                       IF "time_compare"(time_1 := #expire_date_time, time_2 := #current_time, difference_treshold := LT#0s) = true THEN

                           #shaker_batch_code_str[#runtime_shaker_index_finding_Instance.shaker_index - 1] := #batch_no;

                           IF #chemical = "DB_chemical_code".Application_bottle_code_Primer_DV954V1 THEN
                               #shaker_chemical_type_str[#runtime_shaker_index_finding_Instance.shaker_index - 1] := 'Primer DV 954 V1';
                               #shaker_door_lock_control_Instance.mixer_door_lock_enable[#runtime_shaker_index_finding_Instance.shaker_index - 1] := true;
                               #label_scanned := false;
                           ELSIF #chemical = "DB_chemical_code".Application_bottle_code_Primer_SIKA_207 THEN
                               #shaker_chemical_type_str[4] := 'Primer SIKA 207';
                               #shaker_door_lock_control_Instance.mixer_door_lock_enable[4] := true;
                               #label_scanned := false;
                           ELSE
                               #error_state := 256;
                               #shake_deinit := true;
                               #shaker_batch_code_str[#runtime_shaker_index_finding_Instance.shaker_index - 1] := '';
                               #shaker_chemical_type_str[#runtime_shaker_index_finding_Instance.shaker_index - 1] := '';
                           END_IF;
                       ELSE
                           #error_state := 8;
                           #shake_deinit := true;
                           #shaker_batch_code_str[#runtime_shaker_index_finding_Instance.shaker_index - 1] := '';
                           #shaker_chemical_type_str[#runtime_shaker_index_finding_Instance.shaker_index - 1] := '';
                       END_IF;
                   ELSE
                       #error_state := 128;
                       #shake_deinit := true;
                       #shaker_batch_code_str[#runtime_shaker_index_finding_Instance.shaker_index - 1] := '';
                       #shaker_chemical_type_str[#runtime_shaker_index_finding_Instance.shaker_index - 1] := '';
                   END_IF;
               END_IF;
           ELSE
               #error_state := 4;
               #shake_deinit := true;
           END_IF;

       END_IF;
       (* shaking procedure terminated *)
       IF #shaker_index_pre > 0 AND #runtime_shaker_index_finding_Instance.shaker_index = 0 THEN
           #shake_deinit := true;
       END_IF;

       #shaker_index_pre := #runtime_shaker_index_finding_Instance.shaker_index;
   END_IF;

   IF #shake_deinit = true THEN
       #runtime_shaker_index_finding_Instance.shaker_index := 0;
       #shake_deinit := false;
       #label_scanned := false;
       #shaking_enable := false;
       #hmi_label_index := 0;
   END_IF;

   (* hmi info label shaking *)
   #runtime_shake_count_expiration_Instance(mixer_1_presence_sensor_1:=#shaker_1_door_1_bottle_presence,
                                            mixer_1_presence_sensor_2:=#shaker_1_door_2_bottle_presence,
                                            mixer_2_presence_sensor_1:=#shaker_2_door_1_bottle_presence,
                                            mixer_2_presence_sensor_2:=#shaker_2_door_2_bottle_presence,
                                            mixer_3_presence_sensor_1:=#shaker_3_door_1_bottle_presence,
                                            primer_DV954V1_shake_time:=#primer_DV954V1_shake_time,
                                            primer_SIKA_207_shake_time:=#primer_SIKA_207_shake_time,
                                            fs_mixer_door_lock_enable:=#shaker_door_lock_control_Instance.mixer_door_lock_enable,
                                            fs_shaker_chemical_type_str:=#shaker_chemical_type_str,
                                            fs_shaker_batch_code_str:=#shaker_batch_code_str);


   #shaker_door_lock_control_Instance(mixer_1_door_1_lock := #shaker_1_door_1_lock,
                                      mixer_1_door_2_lock := #shaker_1_door_2_lock,
                                      mixer_2_door_1_lock := #shaker_2_door_1_lock,
                                      mixer_2_door_2_lock := #shaker_2_door_2_lock,
                                      mixer_3_door_1_lock := #shaker_3_door_1_lock,
                                      mixer_1_door_1_is_close := #shaker_1_door_1_position,
                                      mixer_1_door_2_is_close := #shaker_1_door_2_position,
                                      mixer_2_door_1_is_close := #shaker_2_door_1_position,
                                      mixer_2_door_2_is_close := #shaker_2_door_2_position,
                                      mixer_3_door_1_is_close := #shaker_3_door_1_position,
                                      mixer_1_presence_sensor_1 := #shaker_1_door_1_bottle_presence,
                                      mixer_1_presence_sensor_2 := #shaker_1_door_2_bottle_presence,
                                      mixer_2_presence_sensor_1 := #shaker_2_door_1_bottle_presence,
                                      mixer_2_presence_sensor_2 := #shaker_2_door_2_bottle_presence,
                                      mixer_3_presence_sensor_1 := #shaker_3_door_1_bottle_presence);
END_FUNCTION_BLOCK

FUNCTION_BLOCK "runtime_shaker_index_finding"   // FB25, SCL
{ S7_Optimized_Access := 'FALSE' }
VERSION : 0.1
BEGIN
   IF #shaker_index > 0 THEN
       IF ((#mixer_1_bottle_1_pre = false AND #mixer_1_presence_sensor_1 = true) OR
           (#mixer_1_bottle_2_pre = false AND #mixer_1_presence_sensor_2 = true) OR
           (#mixer_2_bottle_1_pre = false AND #mixer_2_presence_sensor_1 = true) OR
           (#mixer_2_bottle_2_pre= false AND #mixer_2_presence_sensor_2 = true) OR
           (#mixer_3_bottle_1_pre = false AND #mixer_3_presence_sensor_1 = true)) THEN
           #shaker_index := 0;
           #error_state_identifier := 4096;
       ELSIF ((#mixer_1_bottle_1_pre = true AND #mixer_1_presence_sensor_1 = false) OR
           (#mixer_1_bottle_2_pre = true AND #mixer_1_presence_sensor_2 = false) OR
           (#mixer_2_bottle_1_pre = true AND #mixer_2_presence_sensor_1 = false) OR
           (#mixer_2_bottle_2_pre = true AND #mixer_2_presence_sensor_2 = false) OR
           (#mixer_3_bottle_1_pre = true AND #mixer_3_presence_sensor_1 = false)) THEN
           #shaker_index := 0;
       END_IF;
   ELSE
       IF #mixer_1_bottle_1_pre = false AND #mixer_1_presence_sensor_1 = true THEN
           #shaker_index := 1;
       ELSIF #mixer_1_bottle_2_pre = false AND #mixer_1_presence_sensor_2 = true THEN
           #shaker_index := 2;
       ELSIF #mixer_2_bottle_1_pre = false AND #mixer_2_presence_sensor_1 = true THEN
           #shaker_index := 3;
           #shaking_enable := true;
       ELSIF #mixer_2_bottle_2_pre = false AND #mixer_2_presence_sensor_2 = true THEN
           #shaker_index := 4;
       ELSIF #mixer_3_bottle_1_pre = false AND #mixer_3_presence_sensor_1 = true THEN
           #shaker_index := 5;
       END_IF;

       IF #shaker_index > 0 THEN
           #shaking_enable := true;
       END_IF;
   END_IF;

   #mixer_1_bottle_1_pre := #mixer_1_presence_sensor_1;
   #mixer_1_bottle_2_pre := #mixer_1_presence_sensor_2;
   #mixer_2_bottle_1_pre := #mixer_2_presence_sensor_1;
   #mixer_2_bottle_2_pre := #mixer_2_presence_sensor_2;
   #mixer_3_bottle_1_pre := #mixer_3_presence_sensor_1;
END_FUNCTION_BLOCK

FUNCTION_BLOCK "runtime_shake_count_expiration"   // FB26, SCL
{ S7_Optimized_Access := 'FALSE' }
VERSION : 0.1
BEGIN
   (* shaking time expiration *)
   IF ("Clock_1Hz" = true AND #clock_pre = false) THEN
       IF RD_SYS_T(#current_date_time) < 2 THEN
           #index := 0;
           WHILE #index < 5 DO
               IF #fs_mixer_door_lock_enable[#index] = true THEN
                   IF #fs_shaker_chemical_type_str[#index] = 'Primer DV 954 V1' THEN
                       #mixer_expiration_sec[#index] := LINT_TO_INT(TIME_TO_LINT(#primer_DV954V1_shake_time) / 1000) - DINT_TO_INT(TIME_TO_DINT(T_DIFF(IN2 := #fs_mixer_expiration[#index], IN1 := #current_date_time)) / 1000);
                   ELSIF #fs_shaker_chemical_type_str[#index] = 'Primer SIKA 207' THEN
                       #mixer_expiration_sec[#index] := LINT_TO_INT(TIME_TO_LINT(#primer_SIKA_207_shake_time) / 1000) - DINT_TO_INT(TIME_TO_DINT(T_DIFF(IN2 := #fs_mixer_expiration[#index], IN1 := #current_date_time)) / 1000);
                   END_IF;
               ELSE
                   #mixer_expiration_sec[#index] := 0;
                   #fs_shaker_expiration_str[#index] := '0s';
               END_IF;

               (*nastavit příznak protřepání*)
               IF #mixer_expiration_sec[#index] = 1 THEN
                   #bottle_shaked[#index] := true;
               END_IF;

               IF #mixer_expiration_sec[#index] <= 0 THEN
                   #fs_mixer_door_lock_enable[#index] := false;
               ELSE
                   #temp_string := '    ';
                   IF #mixer_expiration_sec[#index] >= 100 THEN
                       #temp_string[4] := 's';
                       #temp_string[3] := ((#mixer_expiration_sec[#index] MOD 10)) + 48;
                       #temp_string[2] := ((#mixer_expiration_sec[#index] MOD 100 / 10) MOD 10) + 48;
                       #temp_string[1] := (#mixer_expiration_sec[#index] / 100) + 48;
                   ELSIF #mixer_expiration_sec[#index] >= 10 AND #mixer_expiration_sec[#index] < 100 THEN
                       #temp_string[3] := 's';
                       #temp_string[2] := ((#mixer_expiration_sec[#index] MOD 10)) + 48;
                       #temp_string[1] := ((#mixer_expiration_sec[#index]) / 10) + 48;

                   ELSIF #mixer_expiration_sec[#index] < 10 THEN
                       #temp_string[2] := 's';
                       #temp_string[1] := ((#mixer_expiration_sec[#index] MOD 10)) + 48;
                   END_IF;
                   #fs_shaker_expiration_str[#index] := #temp_string;
               END_IF;
               #index := #index + 1;
           END_WHILE;
       END_IF;
   END_IF;

   #clock_pre := "Clock_1Hz";


   (*odeslat informace o protřepání do databáze*)
   IF RD_SYS_T(#current_date_time) < 2 THEN
       ;
   END_IF;
   #expire_date_time_string := CONCAT(IN1 := #expire_date_time_string, IN2 := "copyAndFill"(characterFill := '0', charReplace := '+', stringIn := (DELETE(IN := INT_TO_STRING(#current_date_time.DAY), L := 1, P := 1)), P := 0, char_number := 2));
   #expire_date_time_string := CONCAT(IN1 := #expire_date_time_string, IN2 := '.');
   #expire_date_time_string := CONCAT(IN1 := #expire_date_time_string, IN2 := "copyAndFill"(characterFill := '0', charReplace := '+', stringIn := (DELETE(IN := INT_TO_STRING(#current_date_time.MONTH), L := 1, P := 1)), P := 0, char_number := 2));
   #expire_date_time_string := CONCAT(IN1 := #expire_date_time_string, IN2 := '.');
   #expire_date_time_string := CONCAT(IN1 := #expire_date_time_string, IN2 := "copyAndFill"(characterFill := '0', charReplace := '+', stringIn := (DELETE(IN := UINT_TO_STRING(#current_date_time.YEAR), L := 1, P := 1)), P := 0, char_number := 4));
   #expire_date_time_string := CONCAT(IN1 := #expire_date_time_string, IN2 := '*');
   //time formating
   #expire_date_time_string := CONCAT(IN1 := #expire_date_time_string, IN2 := "copyAndFill"(characterFill := '0', charReplace := '+', stringIn := (DELETE(IN := INT_TO_STRING(#current_date_time.HOUR), L := 1, P := 1)), P := 0, char_number := 2));
   #expire_date_time_string := CONCAT(IN1 := #expire_date_time_string, IN2 := ':');
   #expire_date_time_string := CONCAT(IN1 := #expire_date_time_string, IN2 := "copyAndFill"(characterFill := '0', charReplace := '+', stringIn := (DELETE(IN := INT_TO_STRING(#current_date_time.MINUTE), L := 1, P := 1)), P := 0, char_number := 2));


   IF #bottle_shaked[0] AND #mixer_1_presence_sensor_1 = false THEN
       #database_command_done := "set_table_record_item"(table := 'suplier_bottle',
                                                         record := 'batch_code',
                                                         record_key := #fs_shaker_batch_code_str[0],
                                                         item := 'last_shake',
                                                         new_item_data := #expire_date_time_string,
                                                         server_connection := "tcp_datablock".tcp_connection,
                                                         index := "tcp_datablock".fs_shaker_1_index);

       IF #database_command_done = true THEN
           #bottle_shaked[0] := false;
           #fs_shaker_batch_code_str[0] := '';
           #fs_shaker_chemical_type_str[0] := '';
       END_IF;

   END_IF;

   IF #bottle_shaked[1] AND #mixer_1_presence_sensor_2 = false THEN
       #database_command_done := "set_table_record_item"(table := 'suplier_bottle',
                                                         record := 'batch_code',
                                                         record_key := #fs_shaker_batch_code_str[1],
                                                         item := 'last_shake',
                                                         new_item_data := #expire_date_time_string,
                                                         server_connection := "tcp_datablock".tcp_connection,
                                                         index := "tcp_datablock".fs_shaker_2_index);

       IF #database_command_done = true THEN
           #bottle_shaked[1] := false;
           #fs_shaker_batch_code_str[1] := '';
           #fs_shaker_chemical_type_str[1] := '';
       END_IF;
   END_IF;

   IF #bottle_shaked[2] AND #mixer_2_presence_sensor_1 = false THEN
       #database_command_done := "set_table_record_item"(table := 'suplier_bottle',
                                                         record := 'batch_code',
                                                         record_key := #fs_shaker_batch_code_str[2],
                                                         item := 'last_shake',
                                                         new_item_data := #expire_date_time_string,
                                                         server_connection := "tcp_datablock".tcp_connection,
                                                         index := "tcp_datablock".fs_shaker_3_index);

       IF #database_command_done = true THEN
           #bottle_shaked[2] := false;
           #fs_shaker_batch_code_str[2] := '';
           #fs_shaker_chemical_type_str[2] := '';
       END_IF;
   END_IF;

   IF #bottle_shaked[3] AND #mixer_2_presence_sensor_2 = false THEN
       #database_command_done := "set_table_record_item"(table := 'suplier_bottle',
                                                         record := 'batch_code',
                                                         record_key := #fs_shaker_batch_code_str[3],
                                                         item := 'last_shake',
                                                         new_item_data := #expire_date_time_string,
                                                         server_connection := "tcp_datablock".tcp_connection,
                                                         index := "tcp_datablock".fs_shaker_4_index);

       IF #database_command_done = true THEN
           #bottle_shaked[3] := false;
           #fs_shaker_batch_code_str[3] := '';
           #fs_shaker_chemical_type_str[3] := '';
       END_IF;
   END_IF;

   IF #bottle_shaked[4] AND #mixer_3_presence_sensor_1 = false THEN
       #database_command_done := "set_table_record_item"(table := 'suplier_bottle',
                                                         record := 'batch_code',
                                                         record_key := #fs_shaker_batch_code_str[4],
                                                         item := 'last_shake',
                                                         new_item_data := #expire_date_time_string,
                                                         server_connection := "tcp_datablock".tcp_connection,
                                                         index := "tcp_datablock".fs_shaker_5_index);

       IF #database_command_done = true THEN
           #bottle_shaked[4] := false;
           #fs_shaker_batch_code_str[4] := '';
           #fs_shaker_chemical_type_str[4] := '';
       END_IF;
   END_IF;
END_FUNCTION_BLOCK

FUNCTION_BLOCK "fce_print_sp_botle_label"   // FB27, SCL
{ S7_Optimized_Access := 'FALSE' }
VERSION : 0.1
BEGIN
END_FUNCTION_BLOCK

FUNCTION_BLOCK "fce_filling"   // FB28, SCL
{ S7_Optimized_Access := 'FALSE' }
VERSION : 0.1
BEGIN
END_FUNCTION_BLOCK

FUNCTION "RPA60_HandlerFunction" : Void   // FC2, SCL
{ S7_Optimized_Access := 'FALSE' }
VERSION : 0.1
BEGIN
END_FUNCTION

FUNCTION "setPosition" : Void   // FC5, SCL
{ S7_Optimized_Access := 'FALSE' }
VERSION : 0.1
BEGIN

   IF #positionSensor = #stateOfPositionSensor THEN
           #setPosition := "lockAxis"(valveNewState := #valveNewState,
                                      valve_error_checking:=#valve_error_check,
                                      valve := #valve,
                                      valvePositionSensor := #valvePositionSensor);
       ELSE
           #setPosition := false;
       END_IF;
END_FUNCTION

FUNCTION "StartStation" : Void   // FC6, SCL
{ S7_Optimized_Access := 'FALSE' }
VERSION : 0.1
BEGIN
   (*
   start of station means set true value to the StationStartControlVariable and switch on the lights, but lights are controled from hmi, 
   so they must be switched on only at start
   *)

   IF #startButton = true AND #StationStartControlVariable = false THEN
       #StationStartControlVariable := true;
       #stationLight := true;
   END_IF;
END_FUNCTION

FUNCTION "RPA10B_Main" : Void   // FC7, SCL
{ S7_Optimized_Access := 'FALSE' }
VERSION : 0.1
BEGIN

   IF "RPA10B_datablock".RPA10B_station_start THEN
       IF NOT "RPA10B_LCD_switch_manual_automat" THEN

           "server_connection_handler"(error_state_lock_identifier := 1000,
                                       fatal_error_state_lock := "RPA10B_datablock".PA10B_fatal_error_state_lock,
                                       database_connection := "tcp_datablock".tcp_connection,
                                       error_state_lock := "RPA10B_datablock".PA10B_error_state_lock);

           (* scanner handler *)
           "RPA10B_Scanner_DB"("PORT" := "PA10B~CM_PtP_1",
                               BUFFER := "RPA10B_Scanner_DB".ReceiveBuffer,
                               NDR => "RPA10B_Scanner_DB".NDR,
                               ERROR => "RPA10B_Scanner_DB".ERROR,
                               STATUS => "RPA10B_Scanner_DB".STATUS,
                               LENGTH => "RPA10B_Scanner_DB".LENGTH);

           IF "RPA10B_Scanner_DB".NDR = true THEN
               Chars_TO_Strg(Chars := "RPA10B_Scanner_DB".ReceiveBuffer,
                             pChars := 0,
                             Cnt := "RPA10B_Scanner_DB".received_length - 1,
                             Strg => "RPA10B_datablock".RPA10B_scanned_data );
           END_IF;


           "RPA10B_handler_function"();

           "beaconStateControl"(big_fail_state_lock:="RPA10B_datablock".PA10B_big_fail_state_lock,
                                fail_state_lock:="RPA10B_datablock".PA10B_fail_state_lock,
                                error_state_lock:="RPA10B_datablock".PA10B_error_state_lock,
                                fatal_error_state_lock:="RPA10B_datablock".PA10B_fatal_error_state_lock,
                                beaconGreen:="RPA10B_LCD_beacon_green",
                                beaconOrange:="RPA10B_LCD_beacon_orange",
                                beaconRed:="RPA10B_LCD_beacon_red");

           "beaconStateControl"(big_fail_state_lock := "RPA10B_datablock".PA10B_big_fail_state_lock,
                                fail_state_lock := "RPA10B_datablock".PA10B_fail_state_lock,
                                error_state_lock := "RPA10B_datablock".PA10B_error_state_lock,
                                fatal_error_state_lock := "RPA10B_datablock".PA10B_fatal_error_state_lock,
                                beaconGreen := "RPA10B_primerbox_beacon_green",
                                beaconOrange := "RPA10B_primerbox_beacon_orange",
                                beaconRed := "RPA10B_primerbox_beacon_red");

           "sirenPulsingHandler"(fatal_error:="RPA10B_datablock".PA10B_fatal_error_state_lock,
                                 big_fail:="RPA10B_datablock".PA10B_big_fail_state_lock,
                                 siren_handler_enable:="RPA10B_datablock".RPA10B_siren_hadler_enable,
                                 siren:="RPA10B_LCD_beacon_siren");

           "sirenPulsingHandler"(fatal_error := "RPA10B_datablock".PA10B_fatal_error_state_lock,
                                 big_fail := "RPA10B_datablock".PA10B_big_fail_state_lock,
                                 siren_handler_enable:="RPA10B_datablock".RPA10B_siren_hadler_enable,
                                 siren := "RPA10B_primerbox_beacon_siren");

           "bottleLightControl"(bottleInUsage:="RPA10B_datablock".PA10B_bottle_1_usage,
                                stationWorkCyclusState:="RPA10B_datablock".RPA10B_station_work_cyclus_state,
                                bigFailStateLock:="RPA10B_datablock".PA10B_big_fail_state_lock,
                                ErrorStateLock:="RPA10B_datablock".PA10B_error_state_lock,
                                FatalErrorStateLock:="RPA10B_datablock".PA10B_fatal_error_state_lock,
                                sectionFailIdentifier:=203,
                                bottlePresenceSensor:="RPA10B_primerbox_bottle_1",
                                bottle_taking:="RPA10B_datablock".PA10B_bottle_taking,
                                bottleLight:="RPA10B_primerbox_LED_green_bottle_1",
                                failStateLock:="RPA10B_datablock".PA10B_fail_state_lock,
                                buttonConfirmLED:="RPA10B_LCD_LED_blue_confirm_button");

           "bottleLightControl"(bottleInUsage := "RPA10B_datablock".PA10B_bottle_2_usage,
                                stationWorkCyclusState := "RPA10B_datablock".RPA10B_station_work_cyclus_state,
                                bigFailStateLock := "RPA10B_datablock".PA10B_big_fail_state_lock,
                                ErrorStateLock := "RPA10B_datablock".PA10B_error_state_lock,
                                FatalErrorStateLock := "RPA10B_datablock".PA10B_fatal_error_state_lock,
                                sectionFailIdentifier := 204,
                                bottlePresenceSensor := "RPA10B_primerbox_bottle_2",
                                bottle_taking := "RPA10B_datablock".PA10B_bottle_taking,
                                bottleLight := "RPA10B_primerbox_LED_green_bottle_2",
                                failStateLock := "RPA10B_datablock".PA10B_fail_state_lock,
                                buttonConfirmLED := "RPA10B_LCD_LED_blue_confirm_button");

           "feltLightControl"(feltPresenceSensor:="RPA10B_primerbox_felt_presence_sensor",
                              bigFailStateLock:="RPA10B_datablock".PA10B_big_fail_state_lock,
                              ErrorStateLock:="RPA10B_datablock".PA10B_error_state_lock,
                              FatalErrorStateLock:="RPA10B_datablock".PA10B_fatal_error_state_lock,
                              failStateLockIdentifier:=150,
                              feltLED:="RPA10B_primerbox_LED_green_felt",
                              readyLED:="RPA10B_primerbox_LED_green_ready",
                              failStateLock:= "RPA10B_datablock".PA10B_fail_state_lock,
                              notReady:="RPA10B_primerbox_LED_red_NOT_READY",
                              confirmButtonLED:="RPA10B_LCD_LED_blue_confirm_button");
           (*
           "valveErrorHandler"(valveLock:="RPA10B_EJ_1_vacuum_control",
                               valveLockState:="RPA10B_blend_1_vacuum_fix_sensor",
                               valveErrorCheckingState:="RPA10B_datablock".RPA10B_vacuum_R_check_state,
                               fatalErrorSectionLock:=245,
                               confirmButton:="RPA10B_LCD_button_confirm",
                               fatalErrorLock:="RPA10B_datablock".PA10B_fatal_error_state_lock,
                               confirmButtonLED:="RPA10B_LCD_LED_blue_confirm_button");
                               *)
           (*
           "valveErrorHandler"(valveLock := "RPA10B_EJ_2_vacuum_control",
                               valveLockState := "RPA10B_blend_2_vacuum_fix_sensor",
                               valveErrorCheckingState := "RPA10B_datablock".RPA10B_vacuum_L_check_state,
                               fatalErrorSectionLock := 245,
                               confirmButton := "RPA10B_LCD_button_confirm",
                               fatalErrorLock := "RPA10B_datablock".PA10B_fatal_error_state_lock,
                               confirmButtonLED := "RPA10B_LCD_LED_blue_confirm_button");

           "valveErrorHandler"(valveLock := "RPA10B_,
                               valveLockState := "RPA10B_blend_2_vacuum_fix_sensor",
                               valveErrorCheckingState := "RPA10B_datablock".RPA10B_vacuum_L_check_state,
                               fatalErrorSectionLock := 245,
                               confirmButton := "RPA10B_LCD_button_confirm",
                               fatalErrorLock := "RPA10B_datablock".PA10B_fatal_error_state_lock,
                               confirmButtonLED := "RPA10B_LCD_LED_blue_confirm_button");



           *)

           "RPA10B_idler_presence_handler"(errorStateLock := "RPA10B_datablock".PA10B_error_state_lock,
                                           fatalErrorStateLock := "RPA10B_datablock".PA10B_fatal_error_state_lock,
                                           idler_presence_sensor := "RPA10B_idler_presence_sensor",
                                           idler_in_use := "RPA10B_datablock".RPA10B_idler_in_use,
                                           idler_taking := "RPA10B_datablock".RPA10B_idler_taking,
                                           bigFailStateIdentifire := 205,
                                           confirmButton := "RPA10B_LCD_button_confirm",
                                           confirmButtonLed := "RPA10B_LCD_LED_blue_confirm_button",
                                           bigFailStateLock := "RPA10B_datablock".PA10B_big_fail_state_lock);

           IF ("RPA10B_datablock".PA10B_fail_state_lock + "RPA10B_datablock".PA10B_big_fail_state_lock + "RPA10B_datablock".PA10B_error_state_lock + "RPA10B_datablock".PA10B_fatal_error_state_lock) = 0 THEN

               "pa10b_vacuum_cleaner_controll_DB"(vacuum_sensor := "RPA10B_vacuum_sensor",
                                                  vacuum_control_variable := "RPA10B_vacuum_cleaner_switch");
           END_IF;
       END_IF;
   ELSE

       "RPA10B_datablock".RPA10B_idler_in_use := false;
       "RPA10B_datablock".RPA10B_idler_taking := false;
       "RPA10B_datablock".PA10B_bottle_2_usage := false;
       "RPA10B_datablock".PA10B_bottle_1_usage := false;
       "RPA10B_datablock".PA10B_bottle_taking := false;

       "RPA10B_LCD_beacon_green" := false;
       "RPA10B_LCD_beacon_red" := false;
       "RPA10B_LCD_beacon_orange" := false;
       "RPA10B_LCD_beacon_siren" := false;
       "RPA10B_primerbox_beacon_green" := false;
       "RPA10B_primerbox_beacon_orange" := false;
       "RPA10B_primerbox_beacon_red" := false;
       "RPA10B_primerbox_beacon_siren" := false;

       "RPA10B_primerbox_LED_green_ready" := false;
       "RPA10B_primerbox_LED_green_felt" := false;
       "RPA10B_primerbox_LED_green_bottle_1" := false;
       "RPA10B_primerbox_LED_green_bottle_2" := false;
       "RPA10B_primerbox_LED_red_NOT_READY" := false;
       "RPA10B_primerbox_LED_orange_change_pad" := false;
       "RPA10B_LCD_LED_blue_confirm_button" := false;

       "RPA10B_vavle_aretation_unlock" := true;
       "RPA10B_vavle_aretation_lock" := false;

       "RPA10B_vavle_seal_idler_unlock" := true;
       "RPA10B_vavle_seal_idler_lock" := false;

       "RPA10B_datablock".PA10B_big_fail_state_lock := 0;
       "RPA10B_datablock".PA10B_error_state_lock := 0;
       "RPA10B_datablock".PA10B_fail_state_lock := 0;
       "RPA10B_datablock".PA10B_fatal_error_state_lock := 0;

       "RPA10B_datablock".RPA10B_instruction_list_index := 255;

       "RPA10B_EJ_1_vacuum_control" := false;
       "RPA10B_EJ_2_vacuum_control" := false;
       "RPA10B_EJ_1_eject" := "RPA10B_EJ_1_vacuum_sensor";
       "RPA10B_EJ_2_eject" := "RPA10B_EJ_2_vacuum_sensor";

       "RPA10B_datablock".RPA10B_station_work_cyclus_state := "RPA10B_go_to_home_position";
       "RPA10B_light" := false;

       "StartStation"(startButton:="RPA10B_LCD_button_start",
                      StationStartControlVariable:="RPA10B_datablock".RPA10B_station_start,
                      stationLight:="RPA10B_light");

       "startButtonLightControlHandler"(stationActivitycontrolVariable:="RPA10B_datablock".RPA10B_station_start ,
                                        startButtonLED:="RPA10B_LCD_LED_green_start_button");

   END_IF;


   IF "RPA10B_datablock".RPA10B_station_monitoring_send = true THEN
       "RPA10B_datablock".RPA10B_station_monitoring_send := NOT "pa10b_station_monitoring"(fail_state := "RPA10B_datablock".PA10B_fail_state_lock,
                                                                                           big_fail_state := "RPA10B_datablock".PA10B_big_fail_state_lock,
                                                                                           error_state := "RPA10B_datablock".PA10B_error_state_lock,
                                                                                           fatal_error_state := "RPA10B_datablock".PA10B_fatal_error_state_lock,
                                                                                           work_cyclus_state := "RPA10B_datablock".RPA10B_instruction_list_index,
                                                                                           current_left_cover_code := "RPA10B_datablock".RPA10B_left_cover_code,
                                                                                           current_right_cover_code := "RPA10B_datablock".RPA10B_right_cover_code,
                                                                                           station_activity_state := "RPA10B_datablock".RPA10B_station_start,
                                                                                           position_sensor_1 := "RPA10B_code_position_1",
                                                                                           position_sensor_2 := "RPA10B_code_position_2",
                                                                                           server_connection := "tcp_datablock".tcp_connection,
                                                                                           index:="tcp_datablock".pa10b_station_state_index);
   ELSE
       IF "RPA10B_datablock".RPA10B_fail_state_pre <> "RPA10B_datablock".PA10B_fail_state_lock OR
           "RPA10B_datablock".RPA10B_big_fail_state_pre <> "RPA10B_datablock".PA10B_big_fail_state_lock OR 
           "RPA10B_datablock".RPA10B_error_state_pre <> "RPA10B_datablock".PA10B_error_state_lock OR
           "RPA10B_datablock".RPA10B_fata_error_state_pre <> "RPA10B_datablock".PA10B_fatal_error_state_lock OR
           "RPA10B_datablock".RPA10B_work_cyclus_state_pre <> "RPA10B_datablock".RPA10B_instruction_list_index OR
           "RPA10B_datablock".RPA10B_left_cover_code_pre <> "RPA10B_datablock".RPA10B_left_cover_code OR
           "RPA10B_datablock".RPA10B_right_cover_code_pre <> "RPA10B_datablock".RPA10B_right_cover_code OR
           "RPA10B_datablock".RPA10B_station_activity_state_pre <> "RPA10B_datablock".RPA10B_station_start OR
           "RPA10B_datablock".RPA10B_position_sensor_1_pre <> "RPA10B_code_position_1" OR
           "RPA10B_datablock".RPA10B_position_sensor_2_pre <> "RPA10B_code_position_2" THEN
           "RPA10B_datablock".RPA10B_station_monitoring_send := true;
       END_IF;

       "RPA10B_datablock".RPA10B_fail_state_pre := "RPA10B_datablock".PA10B_fail_state_lock;
       "RPA10B_datablock".RPA10B_big_fail_state_pre := "RPA10B_datablock".PA10B_big_fail_state_lock;
       "RPA10B_datablock".RPA10B_error_state_pre := "RPA10B_datablock".PA10B_error_state_lock;
       "RPA10B_datablock".RPA10B_fata_error_state_pre := "RPA10B_datablock".PA10B_fatal_error_state_lock;
       "RPA10B_datablock".RPA10B_work_cyclus_state_pre := "RPA10B_datablock".RPA10B_instruction_list_index;
       "RPA10B_datablock".RPA10B_left_cover_code_pre := "RPA10B_datablock".RPA10B_left_cover_code;
       "RPA10B_datablock".RPA10B_right_cover_code_pre := "RPA10B_datablock".RPA10B_right_cover_code;
       "RPA10B_datablock".RPA10B_station_activity_state_pre := "RPA10B_datablock".RPA10B_station_start;
       "RPA10B_datablock".RPA10B_position_sensor_1_pre := "RPA10B_code_position_1";
       "RPA10B_datablock".RPA10B_position_sensor_2_pre := "RPA10B_code_position_2";
   END_IF;
END_FUNCTION

FUNCTION "RPA30_changePadHandler" : Void   // FC8, SCL
{ S7_Optimized_Access := 'FALSE' }
VERSION : 0.1
BEGIN


   IF "checkFailStateLock"(failStateLock := #failStateLock,
                               bigFailStateLock := #bigFailStateLock,
                               ErrorStateLock := #ErrorStateLock,
                               FatalErrorStateLock := #FatalErrorStateLock,
                               failStatelockIdetifier := #failStatelockIdetifier) THEN


       "RPA30_F_TRIGR_DB"(CLK:=#padSensor);

       #readyLED := "RPA30_F_TRIGR_DB".STATE AND #padIsChangedButton;
       #notReadyLED := NOT #readyLED;

       #RPA30_changePadHandler := #readyLED;

       IF "RPA30_F_TRIGR_DB".STATE THEN
           #changePedLED := "Clock_0.5Hz";
           IF #padIsChangedButton THEN

               "setOKState"(confirm := true,
                            identifier := #failStatelockIdetifier,
                            confirm_blinking := false,
                            blinkConfirmButton => #confirmButtonLED,
                            stateLock := #failStateLock);
               "RPA30_F_TRIGR_DB".STATE := false;
               #changePedLED := false;
           END_IF;
       ELSE
           #RPA30_changePadHandler := false;
           #changePedLED := #notReadyLED;
           IF "setFailState"(identifier := #failStatelockIdetifier,
                                 failStateLock := #failStateLock) THEN
               ;
           END_IF;
       END_IF;

   ELSE
       #RPA30_changePadHandler := false;
   END_IF;
END_FUNCTION

FUNCTION "IFM_StaticApplicationSwitch" : Void   // FC9, SCL
{ S7_Optimized_Access := 'FALSE' }
VERSION : 0.1
BEGIN

   CASE #ApplicationIndex OF
      1:  // Statement section case 1
          #IFM_Input_1 := false;
          #IFM_Intput_2 := false;
      2:  // Statement section case 2 to 4
          #IFM_Input_1 := true;
          #IFM_Intput_2 := false;
       3:
           #IFM_Input_1 := false;
           #IFM_Intput_2 := true;
       4:
           #IFM_Input_1 := true;
           #IFM_Intput_2 := true;
       ELSE  // Statement section ELSE
           #IFM_Input_1 := false;
           #IFM_Intput_2 := false;
   END_CASE;
END_FUNCTION

FUNCTION "beaconStateControl" : Void   // FC11, SCL
{ S7_Optimized_Access := 'FALSE' }
VERSION : 0.1
BEGIN

   // OK state
   IF (#fail_state_lock + #big_fail_state_lock + #error_state_lock + #fatal_error_state_lock) = 0 THEN
       #beaconGreen := true;
       #beaconOrange := false;
       #beaconRed := false;
   ELSE
       IF (#error_state_lock + #fatal_error_state_lock) > 0 THEN
           #beaconGreen := false;
           #beaconOrange := false;
           #beaconRed := true;
       ELSE
           IF (#fail_state_lock + #big_fail_state_lock) > 0 THEN
               #beaconGreen := false;
               #beaconOrange := true;
               #beaconRed := false;
           END_IF;
       END_IF;
   END_IF;
   // fail/big fail state



   (*
   CASE #stateControlVariable OF
       0:  // OK
           #beaconGreen := true;
           #beaconOrange := false;
           #beaconRed := false;
       1,2: // fail/bad fail
           #beaconGreen := false;
           #beaconOrange := true;
           #beaconRed := false;
       3,4: //error/ fatal error
           #beaconGreen := false;
           #beaconOrange := false;
           #beaconRed := true;
       ELSE  // undefined state
           #beaconGreen := true;
           #beaconOrange := true;
           #beaconRed := true;
   END_CASE;

   *)
END_FUNCTION

FUNCTION "checkFailStateLock" : Void   // FC12, SCL
{ S7_Optimized_Access := 'FALSE' }
VERSION : 0.1
BEGIN

   IF #bigFailStateLock = 0 AND #ErrorStateLock = 0 AND #FatalErrorStateLock = 0 THEN
       IF #failStateLock = 0 OR #failStateLock = #failStatelockIdetifier THEN
           #checkFailStateLock := true;
       ELSE
           #checkFailStateLock := false;
       END_IF;
   ELSE
       #checkFailStateLock := false;
   END_IF;
END_FUNCTION

FUNCTION "checkBigFailStateLock" : Void   // FC13, SCL
{ S7_Optimized_Access := 'FALSE' }
VERSION : 0.1
BEGIN

   IF #ErrorStateLock = 0 AND #FatalErrorStateLock = 0 THEN
       IF #badFailStateLock = 0 OR #badFailStateLock = #badFailStatelockIdetifier THEN
           #checkBigFailStateLock := true;
       ELSE
           #checkBigFailStateLock := false;
       END_IF;
   ELSE
       #checkBigFailStateLock := false;
   END_IF;
END_FUNCTION

FUNCTION "checkErrorStateLock" : Void   // FC14, SCL
{ S7_Optimized_Access := 'FALSE' }
VERSION : 0.1
BEGIN

   IF #FatalErrorStateLock = 0 THEN
       IF #ErrorStateLock = 0 OR #ErrorStateLock = #ErrorStatelockIdetifier THEN
           #checkErrorStateLock := true;
       ELSE
           #checkErrorStateLock := false;
       END_IF;
   ELSE
       #checkErrorStateLock := false;
   END_IF;
END_FUNCTION

FUNCTION "checkFatalErrorStateLock" : Void   // FC15, SCL
{ S7_Optimized_Access := 'FALSE' }
VERSION : 0.1
BEGIN

   IF #FatalErrorStateLock = 0 OR #FatalErrorStateLock = #FatalErrorStatelockIdetifier THEN
       #checkFatalErrorStateLock := true;
   ELSE
       #checkFatalErrorStateLock := false;
   END_IF;
END_FUNCTION

FUNCTION "sirenPulsingHandler" : Void   // FC16, SCL
{ S7_Optimized_Access := 'FALSE' }
VERSION : 0.1
BEGIN
   (*
   creat system clock byte
   *)
   IF #siren_handler_enable THEN
       IF #fatal_error = 0 AND #big_fail = 0 THEN
           #siren := false;
       ELSE
           #siren := "Clock_0.5Hz";
       END_IF;
   END_IF;
END_FUNCTION

FUNCTION "setOKState" : Void   // FC17, SCL
{ S7_Optimized_Access := 'FALSE' }
VERSION : 0.1
BEGIN
   (*
   pokud je volžen odkaz na stav tlačítka, pak bude jeho stav false a nastaví se kontrolní proměnná pro zahájení blikání potvrzovacího tlačítka
   pokud se má stav nastavit okamžitě vloží se do funkce hodnota true a dojde k okamžitému nastavení stavu
   *)

   IF #stateLock = #identifier THEN
       IF #confirm = true THEN
           #blinkConfirmButton := false;
           #stateLock := 0;
       ELSE
           #blinkConfirmButton := "Clock_0.5Hz" AND #confirm_blinking;
       END_IF;
   END_IF;
END_FUNCTION

FUNCTION "RPA30_Main" : Void   // FC19, SCL
{ S7_Optimized_Access := 'FALSE' }
VERSION : 0.1
BEGIN
   //main function of station

   IF "RPA30_DataBlock".RPA30_Start = true THEN
       //cyclus handler function

       IF NOT "RPA30R_LCDSwitchAutomat_Manual" THEN

           "server_connection_handler"(error_state_lock_identifier:=1000,
                                       fatal_error_state_lock:="RPA30_DataBlock".RPA30_fatalErrorStateLock,
                                       database_connection:="tcp_datablock".tcp_connection,
                                       error_state_lock:="RPA30_DataBlock".RPA30_ErrorStateLock);

           "RPA30_Scanner_DB"("PORT" := "pa30~CM_PtP_A14_1",
                              BUFFER := "RPA30_Scanner_DB".ReceiveBuffer);

           IF "RPA30R_LCDButtonConfirmSignal" = true THEN
               "RPA30_DataBlock".RPA30_ErrorStateLock := 0;
               "RPA30_DataBlock".RPA30_fatalErrorStateLock := 0;
               "RPA30_DataBlock".RPA30_fail_state_pre := 0;
               "RPA30_DataBlock".RPA30_bigFailStateLock := 0;
           END_IF;

           IF "RPA30_Scanner_DB".NDR = true THEN
               Chars_TO_Strg(Chars := "RPA30_Scanner_DB".ReceiveBuffer,
                             pChars := 0,
                             Cnt := "RPA30_Scanner_DB".LENGTH - 1,
                             Strg => "RPA30_DataBlock".RPA30_scannedData);
           END_IF;

           IF "RPA30_DataBlock".RPA30_fatalErrorStateLock <> 150 AND "RPA30_DataBlock".RPA30_ErrorStateLock <> 155 THEN

               "RPA30_IFM_point_checking_DB"(primerbox_siren := "RPA30R_Beacon_2_PrimerBoxSiren",
                                             execute := "RPA30_DataBlock".ifm_run,
                                             ifm_side := "RPA30_DataBlock".ifm_side,
                                             keyence_enable := ("RPA30_DataBlock".keyence_enable));
           END_IF;

           (* scan bottle of remover when is changed *)
           IF "RPA30_DataBlock".RPA30_remover_bottle_state_pre = false AND "RPA30R_PrimerPA30SensorBottleRemover208" = true THEN
               IF "RPA30_DataBlock".RPA30_ErrorStateLock = 400 OR "RPA30_DataBlock".RPA30_ErrorStateLock = 401 OR "RPA30_DataBlock".RPA30_ErrorStateLock = 402 OR "RPA30_DataBlock".RPA30_ErrorStateLock = 403 THEN
                   "RPA30R_LedBlueConfirm" := "Clock_0.5Hz";
                   IF "RPA30R_LCDButtonConfirmSignal" = true THEN
                       "RPA30_DataBlock".RPA30_ErrorStateLock := 0;
                       "RPA30R_LedBlueConfirm" := false;
                   END_IF;
               END_IF;

               "RPA30_DataBlock".RPA30_actual_instruction_index := "RPA30_hmi_scan_remover_bottle";
               IF "setFailState"(identifier := 33,
                                     failStateLock := "RPA30_DataBlock".RPA30_failStateLock) THEN
                   IF "RPA30_Scanner_DB".NDR = true THEN
                       #bottle_checking_result := "bottle_label_check"(input_data := "RPA30_DataBlock".RPA30_scannedData, chemical_type := 3);
                       IF #bottle_checking_result = 0 THEN
                           "RPA30_DataBlock".RPA30_actualCodeBottleRemover208 := "RPA30_DataBlock".RPA30_scannedData;
                           "RPA30_DataBlock".RPA30_remover_bottle_state_pre := "RPA30R_PrimerPA30SensorBottleRemover208";
                           "setOKState"(confirm := true,
                                        identifier := 33,
                                        confirm_blinking := false,
                                        blinkConfirmButton => "RPA30R_LedBlueConfirm",
                                        stateLock := "RPA30_DataBlock".RPA30_failStateLock);
                           "RPA30R_LedBlueConfirm" := false;
                       ELSIF #bottle_checking_result = 2 THEN
                           "RPA30_DataBlock".RPA30_ErrorStateLock := 400;
                       ELSIF #bottle_checking_result = 3 THEN
                           "RPA30_DataBlock".RPA30_ErrorStateLock := 401;
                       ELSIF #bottle_checking_result = 4 THEN
                           "RPA30_DataBlock".RPA30_ErrorStateLock := 402;
                       ELSIF #bottle_checking_result = 5 THEN
                           "RPA30_DataBlock".RPA30_ErrorStateLock := 403;
                       END_IF;
                   END_IF;
               END_IF;
           ELSE
               (*
               IF "PLC_datablock".stations_configuration = 0 OR "PLC_datablock".stations_configuration = 2 OR "PLC_datablock".stations_configuration = 4 THEN
                   "RPA30_Handler_function_A"();
               ELSIF "PLC_datablock".stations_configuration = 1 OR "PLC_datablock".stations_configuration = 3 THEN
                   "RPA30_Handler_function_B"();
               END_IF;
               *)
               "RPA30_Handler_function_A"();
               "RPA30_DataBlock".RPA30_remover_bottle_state_pre := "RPA30R_PrimerPA30SensorBottleRemover208";
           END_IF;

           //"RPA30_IFM_runtime_switching"();

           //beacon light control
           "beaconStateControl"(big_fail_state_lock:="RPA30_DataBlock".RPA30_bigFailStateLock,
                                fail_state_lock:="RPA30_DataBlock".RPA30_failStateLock,
                                error_state_lock:="RPA30_DataBlock".RPA30_ErrorStateLock,
                                fatal_error_state_lock:="RPA30_DataBlock".RPA30_fatalErrorStateLock,
                                beaconGreen := "RPA30R_Beacon_2_PrimerBoxGreen",
                                beaconOrange := "RPA30R_Beacon_2_PrimerBoxOrange",
                                beaconRed := "RPA30R_Beacon_2_PrimerBoxRed");

           "beaconStateControl"(big_fail_state_lock:="RPA30_DataBlock".RPA30_bigFailStateLock,
                                fail_state_lock:="RPA30_DataBlock".RPA30_failStateLock,
                                error_state_lock:="RPA30_DataBlock".RPA30_ErrorStateLock,
                                fatal_error_state_lock:="RPA30_DataBlock".RPA30_fatalErrorStateLock,
                                beaconGreen := "RPA30R_Beacon_1_LCDPanelGreen",
                                beaconOrange := "RPA30R_Beacon_1_LCDPanelOrange",
                                beaconRed := "RPA30R_Beacon_1_LCDPanelRed");

           //siren control
           "sirenPulsingHandler"(fatal_error:="RPA30_DataBlock".RPA30_fatalErrorStateLock,
                                 big_fail:="RPA30_DataBlock".RPA30_bigFailStateLock,
                                 siren_handler_enable:="RPA30_DataBlock".RPA30_siren_hadler_enable,
                                 siren := "RPA30R_Beacon_1_LCDPanelSiren");

           //light controller control
           //primer bottle SIKA 207
           "bottleLightControl"(bottleInUsage := "RPA30_DataBlock".RPA30_UseInterval_Primer207,
                                stationWorkCyclusState := "RPA30_DataBlock".RPA30_cyclusState,
                                bigFailStateLock := "RPA30_DataBlock".RPA30_bigFailStateLock,
                                ErrorStateLock := "RPA30_DataBlock".RPA30_ErrorStateLock,
                                FatalErrorStateLock := "RPA30_DataBlock".RPA30_fatalErrorStateLock,
                                sectionFailIdentifier := 100,
                                bottlePresenceSensor := "RPA30R_PrimerPA30SensorBottlePrimer207",
                                bottle_taking:= "RPA30_DataBlock".RPA30_bottle_taking,
                                bottleLight := "RPA30R_PrimerPA30GreenPrimer207",
                                failStateLock := "RPA30_DataBlock".RPA30_failStateLock,
                                buttonConfirmLED := "RPA30R_LedBlueConfirm");

           //remover bottle SIKA 208
           "bottleLightControl"(bottleInUsage := "RPA30_DataBlock".RPA30_UseIntervalBottleRemover208,
                                stationWorkCyclusState := "RPA30_DataBlock".RPA30_cyclusState,
                                bigFailStateLock := "RPA30_DataBlock".RPA30_bigFailStateLock,
                                ErrorStateLock := "RPA30_DataBlock".RPA30_ErrorStateLock,
                                FatalErrorStateLock := "RPA30_DataBlock".RPA30_fatalErrorStateLock,
                                sectionFailIdentifier := 110,
                                bottlePresenceSensor := "RPA30R_PrimerPA30SensorBottleRemover208",
                                bottle_taking := "RPA30_DataBlock".RPA30_bottle_taking,
                                bottleLight := "RPA30R_PrimerPA30GreenRemover208",
                                failStateLock := "RPA30_DataBlock".RPA30_failStateLock,
                                buttonConfirmLED := "RPA30R_LedBlueConfirm");

           "feltLightControl"(feltPresenceSensor := "RPA30R_PrimerPA30SensorFeltEmpty",
                              bigFailStateLock := "RPA30_DataBlock".RPA30_bigFailStateLock,
                              ErrorStateLock := "RPA30_DataBlock".RPA30_ErrorStateLock,
                              FatalErrorStateLock := "RPA30_DataBlock".RPA30_fatalErrorStateLock,
                              failStateLockIdentifier := 300,
                              feltLED := "RPA30R_PrimerPA30GreenFelt",
                              readyLED := "RPA30R_PrimerPA30GreenReady",
                              failStateLock := "RPA30_DataBlock".RPA30_failStateLock,
                              notReady := "RPA30R_PrimerPA30RedNotReady",
                              confirmButtonLED := "RPA30R_LedBlueConfirm");
       END_IF;
   ELSE

       IF "lockAxis"(valvePositionSensor := "RPA30R_PositionCylinderSensorLockY",
                         valveNewState := false,
                         valve_error_checking := "RPA30_DataBlock".RPA30_valveYErrorStateCheck, valve := "RPA30R_ValveCylinderYLock") THEN
           "RPA30_DataBlock".RPA30_bigFailStateLock := 0;
           "RPA30_DataBlock".RPA30_ErrorStateLock := 0;
           "RPA30_DataBlock".RPA30_failStateLock := 0;
           "RPA30_DataBlock".RPA30_fatalErrorStateLock := 0;

           "RPA30_DataBlock".RPA30_bottle_taking := false;
           "RPA30_DataBlock".RPA30_show_smile := false;